REGION Network 9
   RUNG wire#powerrail
      { S7_Templates := "SrcType := Real" } LE_Contact(in1 := #"PID Output", in2 := #RangeY)
      Move(in := 0, out1 => #"Range2.Q")
   END_RUNG
   // the same network as SCL:
   IF #"PID Output" <= #RangeY THEN #"Range2.Q" := 0; END_IF;
END_REGION
END_FUNCTION_BLOCK

// folder: 1}Library/Timers

FUNCTION_BLOCK "TimerDisplay"   // FB2, LAD
{ S7_Optimized_Access := 'TRUE' }
VERSION : 0.1
   VAR_INPUT
      ET : DInt;
   END_VAR
   VAR_OUTPUT
      OUT : String;
   END_VAR
   VAR
      RealH : Real;
      RealM : Real;
      RealS : Real;
      RealMS : Real;
      StringH : String;
      StringM : String;
      StringS : String;
      StringMS : String;
      intH : Int;
      intM : Int;
      intS : Int;
      intMS : Int;
      String5 : String;
      String6 : String;
      String7 : String;
      String8 : String;
   END_VAR
   VAR_TEMP
      "dint-tempH" : DInt;
      "dint-tempM" : DInt;
      "dint-tempS" : DInt;
      "dint-tempMS" : DInt;
      "real-tempH" : Real;
      "real-tempM" : Real;
      "real-tempS" : Real;
      "real-tempMS" : Real;
   END_VAR
BEGIN

REGION Network 1: Reminder of H/M/S/MS
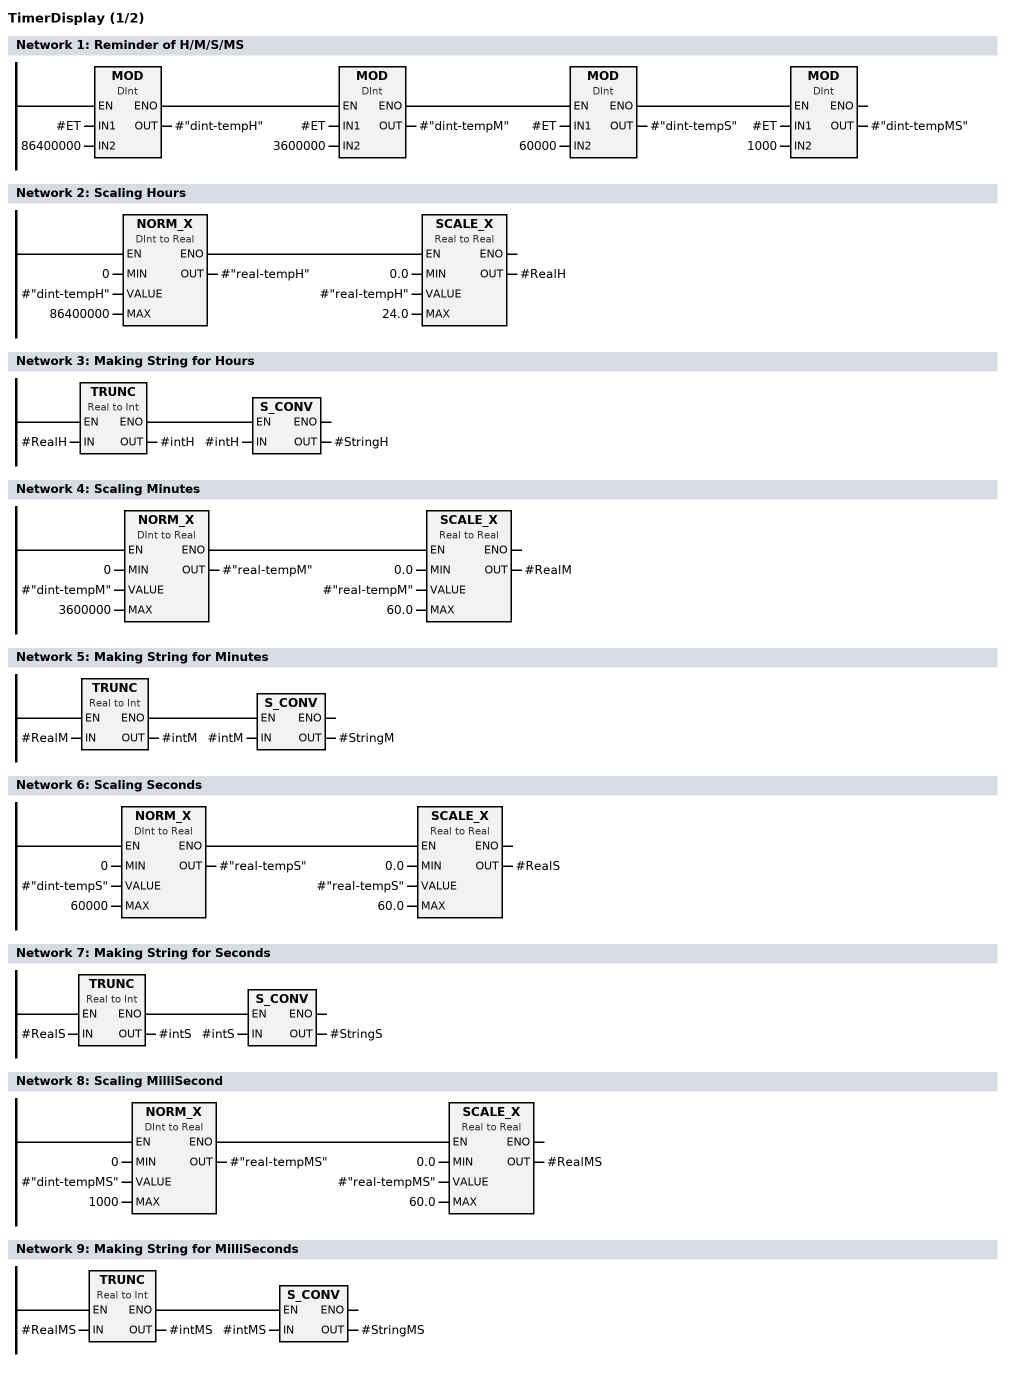
   RUNG wire#powerrail
      { S7_Templates := "SrcType := DInt" } Mod(in1 := #ET, in2 := 86400000, out => #"dint-tempH")
      { S7_Templates := "SrcType := DInt" } Mod(in1 := #ET, in2 := 3600000, out => #"dint-tempM")
      { S7_Templates := "SrcType := DInt" } Mod(in1 := #ET, in2 := 60000, out => #"dint-tempS")
      { S7_Templates := "SrcType := DInt" } Mod(in1 := #ET, in2 := 1000, out => #"dint-tempMS")
   END_RUNG
   // the same network as SCL:
   #"dint-tempH" := #ET MOD 86400000;
   #"dint-tempM" := #ET MOD 3600000;
   #"dint-tempS" := #ET MOD 60000;
   #"dint-tempMS" := #ET MOD 1000;
END_REGION

REGION Network 2: Scaling Hours
   RUNG wire#powerrail
      { S7_Templates := "[SrcType := DInt, DestType := Real]" } Normalize(min := 0, value := #"dint-tempH", max := 86400000, out => #"real-tempH")
      { S7_Templates := "[SrcType := Real, DestType := Real]" } Scale(min := 0.0, value := #"real-tempH", max := 24.0, out => #RealH)
   END_RUNG
   // the same network as SCL:
   #"real-tempH" := NORM_X(MIN := 0, VALUE := #"dint-tempH", MAX := 86400000);
   #RealH := SCALE_X(MIN := 0.0, VALUE := #"real-tempH", MAX := 24.0);
END_REGION

REGION Network 3: Making String for Hours
   #intH := TRUNC(#RealH);
   #StringH := S_CONV(IN := #intH);
END_REGION

REGION Network 4: Scaling Minutes
   RUNG wire#powerrail
      { S7_Templates := "[SrcType := DInt, DestType := Real]" } Normalize(min := 0, value := #"dint-tempM", max := 3600000, out => #"real-tempM")
      { S7_Templates := "[SrcType := Real, DestType := Real]" } Scale(min := 0.0, value := #"real-tempM", max := 60.0, out => #RealM)
   END_RUNG
   // the same network as SCL:
   #"real-tempM" := NORM_X(MIN := 0, VALUE := #"dint-tempM", MAX := 3600000);
   #RealM := SCALE_X(MIN := 0.0, VALUE := #"real-tempM", MAX := 60.0);
END_REGION

REGION Network 5: Making String for Minutes
   #intM := TRUNC(#RealM);
   #StringM := S_CONV(IN := #intM);
END_REGION

REGION Network 6: Scaling Seconds
   RUNG wire#powerrail
      { S7_Templates := "[SrcType := DInt, DestType := Real]" } Normalize(min := 0, value := #"dint-tempS", max := 60000, out => #"real-tempS")
      { S7_Templates := "[SrcType := Real, DestType := Real]" } Scale(min := 0.0, value := #"real-tempS", max := 60.0, out => #RealS)
   END_RUNG
   // the same network as SCL:
   #"real-tempS" := NORM_X(MIN := 0, VALUE := #"dint-tempS", MAX := 60000);
   #RealS := SCALE_X(MIN := 0.0, VALUE := #"real-tempS", MAX := 60.0);
END_REGION

REGION Network 7: Making String for Seconds
   #intS := TRUNC(#RealS);
   #StringS := S_CONV(IN := #intS);
END_REGION

REGION Network 8: Scaling MilliSecond
   RUNG wire#powerrail
      { S7_Templates := "[SrcType := DInt, DestType := Real]" } Normalize(min := 0, value := #"dint-tempMS", max := 1000, out => #"real-tempMS")
      { S7_Templates := "[SrcType := Real, DestType := Real]" } Scale(min := 0.0, value := #"real-tempMS", max := 60.0, out => #RealMS)
   END_RUNG
   // the same network as SCL:
   #"real-tempMS" := NORM_X(MIN := 0, VALUE := #"dint-tempMS", MAX := 1000);
   #RealMS := SCALE_X(MIN := 0.0, VALUE := #"real-tempMS", MAX := 60.0);
END_REGION

REGION Network 9: Making String for MilliSeconds
   #intMS := TRUNC(#RealMS);
   #StringMS := S_CONV(IN := #intMS);
END_REGION

REGION Network 10
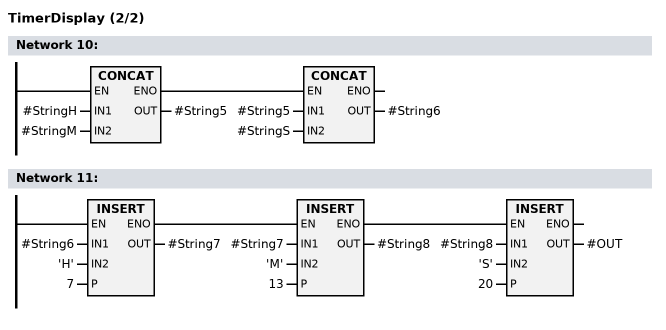
   #String5 := CONCAT(IN1 := #StringH, IN2 := #StringM);
   #String6 := CONCAT(IN1 := #String5, IN2 := #StringS);
END_REGION

REGION Network 11
   #String7 := INSERT(IN1 := #String6, IN2 := 'H', P := 7);
   #String8 := INSERT(IN1 := #String7, IN2 := 'M', P := 13);
   #OUT := INSERT(IN1 := #String8, IN2 := 'S', P := 20);
END_REGION
END_FUNCTION_BLOCK

// folder: 1}Library/Totalizer

FUNCTION_BLOCK "Totalizer_1"   // FB11, LAD
{ S7_Optimized_Access := 'TRUE' }
VERSION : 0.1
   VAR_INPUT
      value : Real;
      interval : Time;
      reset : Bool;
      cycle : Time;
   END_VAR
   VAR_OUTPUT
      Total : Real;
   END_VAR
   VAR
      accum1 : Real;
      accum2 : Real;
      "Timer" : IEC_TIMER;
   END_VAR
   VAR_TEMP
      tempInterval_Real : Real;
      tempInterval_Dint : DInt;
      tempCycle_Real : Real;
      tempCycle_Dint : Real;
      TempCalOne : Real;
      TempCalTwo : Real;
   END_VAR
BEGIN

REGION Network 1 (SCL): Reset Totalizer counts
   IF #reset THEN
       #accum1 := 0.0;
       #accum2 := 0.0;
       RESET_TIMER(#Timer);

   END_IF;
END_REGION

REGION Network 2 (SCL): Convert time into REAL
   #tempInterval_Real := TIME_TO_DINT (#interval);
   #tempCycle_Real := TIME_TO_DINT(#cycle);
END_REGION

REGION Network 3: Calculations for accum1
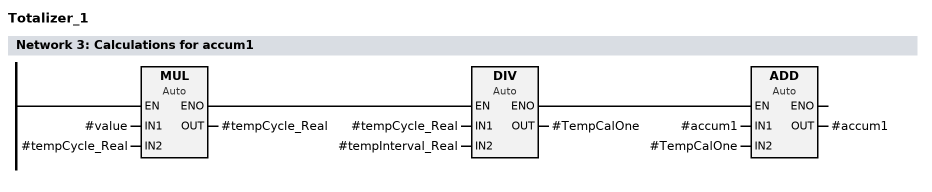
   RUNG wire#powerrail
      Mul(in1 := #value, in2 := #tempCycle_Real, out => #tempCycle_Real)
      Div(in1 := #tempCycle_Real, in2 := #tempInterval_Real, out => #TempCalOne)
      Add(in1 := #accum1, in2 := #TempCalOne, out => #accum1)
   END_RUNG
   // the same network as SCL:
   #tempCycle_Real := #value * #tempCycle_Real;
   #TempCalOne := #tempCycle_Real / #tempInterval_Real;
   #accum1 := #accum1 + #TempCalOne;
END_REGION

REGION Network 4 (SCL): Add the counters and reinitialize accum1
   IF #accum1 >= 1000.0 THEN
       #accum2 := 1000.0 + #accum2;
       #accum1 := 0.0;
   END_IF;

   #Total := #accum1 + #accum2;
END_REGION
END_FUNCTION_BLOCK

FUNCTION_BLOCK "Totalizer"   // FB17, LAD
{ S7_Optimized_Access := 'TRUE' }
VERSION : 0.1
   VAR_INPUT
      value : Real;
      interval : Time;
      reset : Bool;
      cycle : Time;
   END_VAR
   VAR_OUTPUT
      Total : Real;
   END_VAR
   VAR
      accum1 : Real;
      accum2 : Real;
      "Timer" : IEC_TIMER;
   END_VAR
   VAR_TEMP
      tempInterval_Real : Real;
      tempInterval_Dint : DInt;
      tempCycle_Real : Real;
      tempCycle_Dint : Real;
      TempCalOne : Real;
      TempCalTwo : Real;
   END_VAR
BEGIN

REGION Network 1 (SCL): Reset Totalizer counts
   IF #reset THEN
       #accum1 := 0.0;
       #accum2 := 0.0;
       #Total := 0.0;
       RESET_TIMER(#Timer);

   END_IF;
END_REGION

REGION Network 2 (SCL): Convert time into REAL
   #tempInterval_Real := TIME_TO_DINT (#interval);
   #tempCycle_Real := TIME_TO_DINT(#cycle);
END_REGION

REGION Network 3: Calculations for accum1
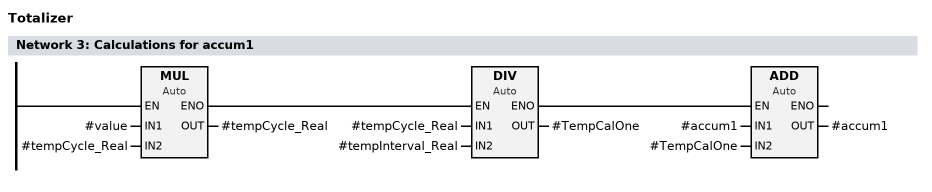
   RUNG wire#powerrail
      Mul(in1 := #value, in2 := #tempCycle_Real, out => #tempCycle_Real)
      Div(in1 := #tempCycle_Real, in2 := #tempInterval_Real, out => #TempCalOne)
      Add(in1 := #accum1, in2 := #TempCalOne, out => #accum1)
   END_RUNG
   // the same network as SCL:
   #tempCycle_Real := #value * #tempCycle_Real;
   #TempCalOne := #tempCycle_Real / #tempInterval_Real;
   #accum1 := #accum1 + #TempCalOne;
END_REGION

REGION Network 4 (SCL): Add the counters and reinitialize accum1
   IF #accum1 >= 1000.0 THEN
       #accum2 := 1000.0 + #accum2;
       #accum1 := 0.0;
   END_IF;

   #Total := #accum1 + #accum2;
END_REGION
END_FUNCTION_BLOCK

// folder: 1}Library/VFD

FUNCTION_BLOCK "VFD_PNCtrl"   // FB9, SCL
TITLE = VFD Controlled by Profinet
{ S7_Optimized_Access := 'TRUE' }
VERSION : 0.1
   VAR_INPUT
      EnableBlock : Bool;
      EnableAxis : Bool;
      AckError : Bool;
      SpeedSP_Perc : Real;   // Speed SP in Percentage 0-100%
      RefSpeed : Real;   // Reference Speed in RPM (parameter p2000)
      ConfigAxis : Word := 16#003F;
      HWIDSTW : Hw_Io;
      HWIDZSW : Hw_Io;
   END_VAR
   VAR_OUTPUT
      AxisEnabled : Bool;
      Lockout : Bool;
      ActVelocity_Perc : Real;
      ActVelocity_RPM : Real;
      Error : Bool;
      Status : Word;
      DiagId : Word;
   END_VAR
   VAR
      SP_Rpm : Real;   // Speed SP in RPM
      SinaSpeed_Instance : SinaSpeed;
   END_VAR
BEGIN
   //******************************************************************************
   //Convert Speed SP from Percentage to RPM

   #SP_Rpm := (#SpeedSP_Perc * #RefSpeed) / 100;

   IF #EnableBlock THEN


       #SinaSpeed_Instance(EnableAxis := #EnableAxis,
                           AckError := #AckError,
                           SpeedSp := #SP_Rpm,
                           RefSpeed := #RefSpeed,
                           ConfigAxis := #ConfigAxis,
                           HWIDSTW := #HWIDSTW,
                           HWIDZSW := #HWIDZSW,
                           AxisEnabled => #AxisEnabled,
                           Lockout => #Lockout,
                           ActVelocity => #ActVelocity_Perc,
                           Error => #Error,
                           Status => #Status,
                           DiagId => #DiagId);

   ELSE

       #SinaSpeed_Instance(EnableAxis := FALSE,
                           AckError :=FALSE,
                           SpeedSp := 0.0,
                           RefSpeed := #RefSpeed,
                           ConfigAxis := #ConfigAxis,
                           HWIDSTW := #HWIDSTW,
                           HWIDZSW := #HWIDZSW,
                           AxisEnabled => #AxisEnabled,
                           Lockout => #Lockout,
                           ActVelocity => #ActVelocity_Perc,
                           Error => #Error,
                           Status => #Status,
                           DiagId => #DiagId);


       #Error := FALSE;

   END_IF;

   #ActVelocity_Perc := (#SinaSpeed_Instance.ActVelocity * 100) / #RefSpeed;
   #ActVelocity_RPM := #SinaSpeed_Instance.ActVelocity;
END_FUNCTION_BLOCK

FUNCTION_BLOCK "VFD_Dumbdown"   // FB812, LAD
{ S7_Optimized_Access := 'TRUE' }
VERSION : 0.7
   VAR_INPUT
      IL : Bool := TRUE;   // Interlock
      PLCCommand : Bool;   // Auto Command to Run (logic from PLC to command motor to run)
      RUN_FEEDBACK : Bool;   // Feedback from the drive indicating that it is running
      VFD_FAULT : Bool;   // Feedback from the drive that it is in Fault
      AUTO_SPEED_P : Word;   // Auto Speed Setpoint Command (logic from PLC to command motor speed) Raw 0-27648
      AUTO_SPEED_R : Real;   // Auto Speed Setpoint Command (logic from PLC to command motor speed) Scale 0-100
      SPEED_FEEDBACK : Int;   // Speed Feedback raw Siganl from the drive
   END_VAR
   VAR_OUTPUT
      RUN_CMD : Bool;
      Stop_CMD : Bool;   // Stop Command
      Start_CMD : Bool;   // Start Command
      RST_CMD : Bool;   // VFD Reset
      VFD_SPEED : Int;   // Command Speed Setpoint to VFD
      VFD_TORQUE : Int;   // Command Torque Setpoint to VFD
   END_VAR
   VAR
      HMI : Struct   // Struct for HMI
         Controls : Struct
            Mode : Int;   // HOA = Auto, 0 = Off, 1 = Manual (HMI Control), 2 = Auto (PLC Control)
            Start : Bool;   // Mode = 1, Start VFD Command
            Stop : Bool;   // Mode = 1, Stop VFD Command
            Reset : Bool;   // VFD Reset Command
            PLCMOHR : Bool;   // PLC Motor Operating Hours Reset
            Speed_Setpoint : Real;   // Speed Setpoint to Drive Real 0-100.0
         END_STRUCT;
         Status : Struct
            HOAStatus : Int;   // HOA Status
            PLC_MOH : Real;
            LMOH : Real;   // Last Motor Operating Hours
            VFDON : Bool;   // VFD On
            VFD_FAULT : Bool;   // VFD is Faulted
            CMD : Bool;   // Commanding VFD to Run
            IL : Bool;   // Interlock Active
            VFD_SPEED : Real;   // VFD Speed Feedback from the drive
            VFD_TORQUE : Real;
         END_STRUCT;
         Config : Struct
            RCPD_SP : Int := 300;
            Start_PT : Time := T#500MS;
            Stop_PT : Time := T#500MS;
         END_STRUCT;
      END_STRUCT;
      Math : Struct
         MOH1 : DInt;
         MOH2 : Real;
         PLCMOH : Real;   // PLC Motor Operating Hours
         LMOH : Real;
      END_STRUCT;
      OS : Struct
         RON : Bool;   // Remote / HMI On
         ROFF : Bool;   // Remote / HMI Off
         HON : Bool;   // Hand/Local On
         Auto : Bool;   // Auto
         PLCMOHR : Bool;
         LMOH1 : Bool;
         LMOH2 : Bool;
         RST : Bool;   // Reset VFD
         Bipolar : Bool;
         MinuteTime : Bool;
         HoursTime : Real;
         Raw_Auto_Speed_Set : Int;
         Unscale_Return : Word;
      END_STRUCT;
      Motor_max_RPM : Real := 100.0;
      START_CMD_TOF : IEC_TIMER;   // Start Semicode
      STOP_CMD_TOF : IEC_TIMER;
      Reset_Hold_Time : IEC_TIMER;
      Motor_Minute_Counter : IEC_TIMER;
      TIMEOUT : IEC_TIMER;
   END_VAR
   VAR_TEMP   // added for the SCL form of the ladder/FBD networks
      _w1 : Bool;
      _w2 : Bool;
   END_VAR
BEGIN

REGION Network 1: Start VFD
   // Main Logic of the FB
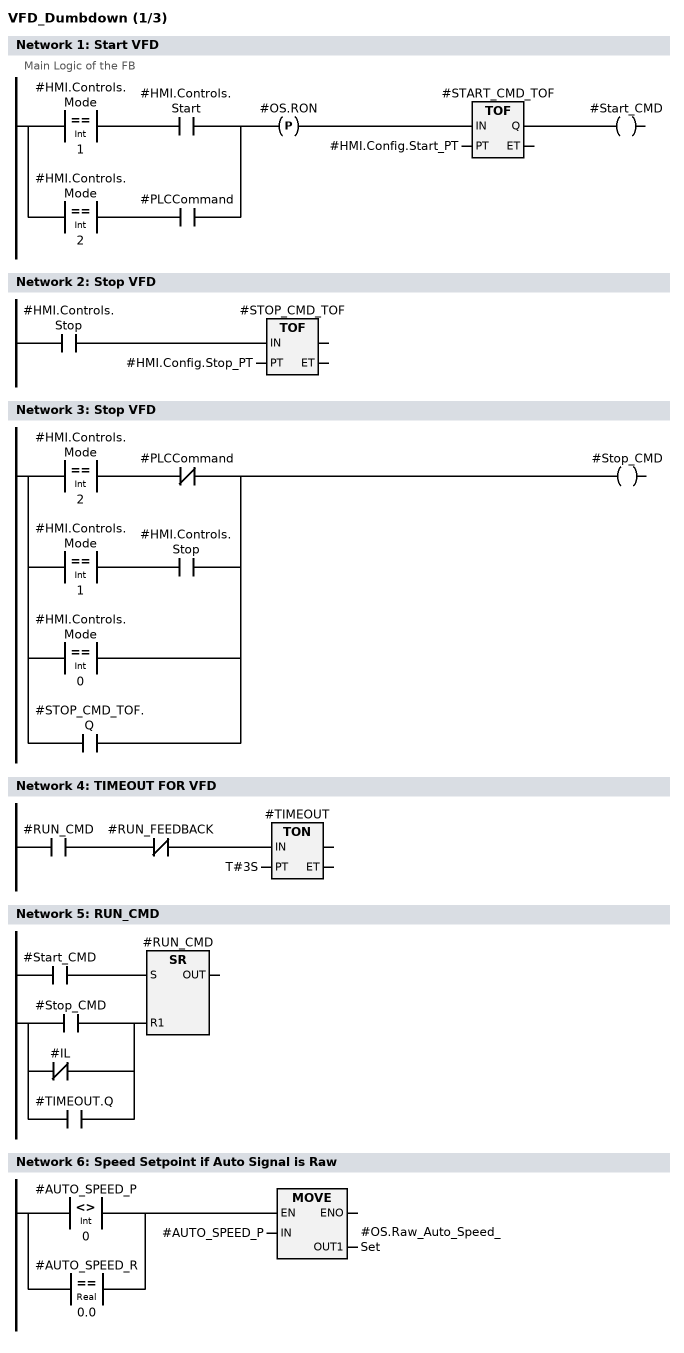
   #_w1 := ((#HMI.Controls.Mode = 1) AND #HMI.Controls.Start) OR ((#HMI.Controls.Mode = 2) AND #PLCCommand);
   #_w2 := #_w1 AND NOT #OS.RON;   // rising edge
   #OS.RON := #_w1;
   #START_CMD_TOF.TOF(IN := #_w2, PT := #HMI.Config.Start_PT);
   #Start_CMD := #START_CMD_TOF.Q;
END_REGION

REGION Network 2: Stop VFD
   #STOP_CMD_TOF.TOF(IN := #HMI.Controls.Stop, PT := #HMI.Config.Stop_PT);
END_REGION

REGION Network 3: Stop VFD
   RUNG wire#powerrail
      { S7_Templates := "SrcType := Int" } EQ_Contact(in1 := #HMI.Controls.Mode, in2 := 2)
      I_Contact( #PLCCommand )
      wire#w1
      Coil( #Stop_CMD )
   END_RUNG
   RUNG wire#powerrail
      { S7_Templates := "SrcType := Int" } EQ_Contact(in1 := #HMI.Controls.Mode, in2 := 1)
      Contact( #HMI.Controls.Stop )
   END_RUNG wire#w1
   RUNG wire#powerrail
      { S7_Templates := "SrcType := Int" } EQ_Contact(in1 := #HMI.Controls.Mode, in2 := 0)
   END_RUNG wire#w1
   RUNG wire#powerrail
      Contact( #STOP_CMD_TOF.Q )
   END_RUNG wire#w1
   // the same network as SCL:
   #Stop_CMD := ((#HMI.Controls.Mode = 2) AND NOT #PLCCommand) OR ((#HMI.Controls.Mode = 1) AND #HMI.Controls.Stop) OR (#HMI.Controls.Mode = 0) OR #STOP_CMD_TOF.Q;
END_REGION

REGION Network 4: TIMEOUT FOR VFD
   #TIMEOUT.TON(IN := #RUN_CMD AND NOT #RUN_FEEDBACK, PT := T#3S);
END_REGION

REGION Network 5: RUN_CMD
   RUNG wire#powerrail
      Contact( #Start_CMD )
      S_SR(operand := #RUN_CMD, r1 := wire#w1)
   END_RUNG
   RUNG wire#powerrail
      Contact( #Stop_CMD )
   END_RUNG wire#w1
   RUNG wire#powerrail
      I_Contact( #IL )
   END_RUNG wire#w1
   RUNG wire#powerrail
      Contact( #TIMEOUT.Q )
   END_RUNG wire#w1
   // the same network as SCL:
   IF #Start_CMD THEN
       #RUN_CMD := TRUE;   // SR flip-flop
   END_IF;
   IF #Stop_CMD OR NOT #IL OR #TIMEOUT.Q THEN #RUN_CMD := FALSE; END_IF;
END_REGION

REGION Network 6: Speed Setpoint if Auto Signal is Raw
   RUNG wire#powerrail
      { S7_Templates := "SrcType := Int" } NE_Contact(in1 := #AUTO_SPEED_P, in2 := 0)
      wire#w1
      { S7_GenerateENO := "TRUE" } Move(in := #AUTO_SPEED_P, out1 => #OS.Raw_Auto_Speed_Set)
   END_RUNG
   RUNG wire#powerrail
      { S7_Templates := "SrcType := Real" } EQ_Contact(in1 := #AUTO_SPEED_R, in2 := 0.0)
   END_RUNG wire#w1
   // the same network as SCL:
   IF (#AUTO_SPEED_P <> 0) OR (#AUTO_SPEED_R = 0.0) THEN #OS.Raw_Auto_Speed_Set := #AUTO_SPEED_P; END_IF;
END_REGION

REGION Network 7: Speed Setpoint if Auto Signal is Real
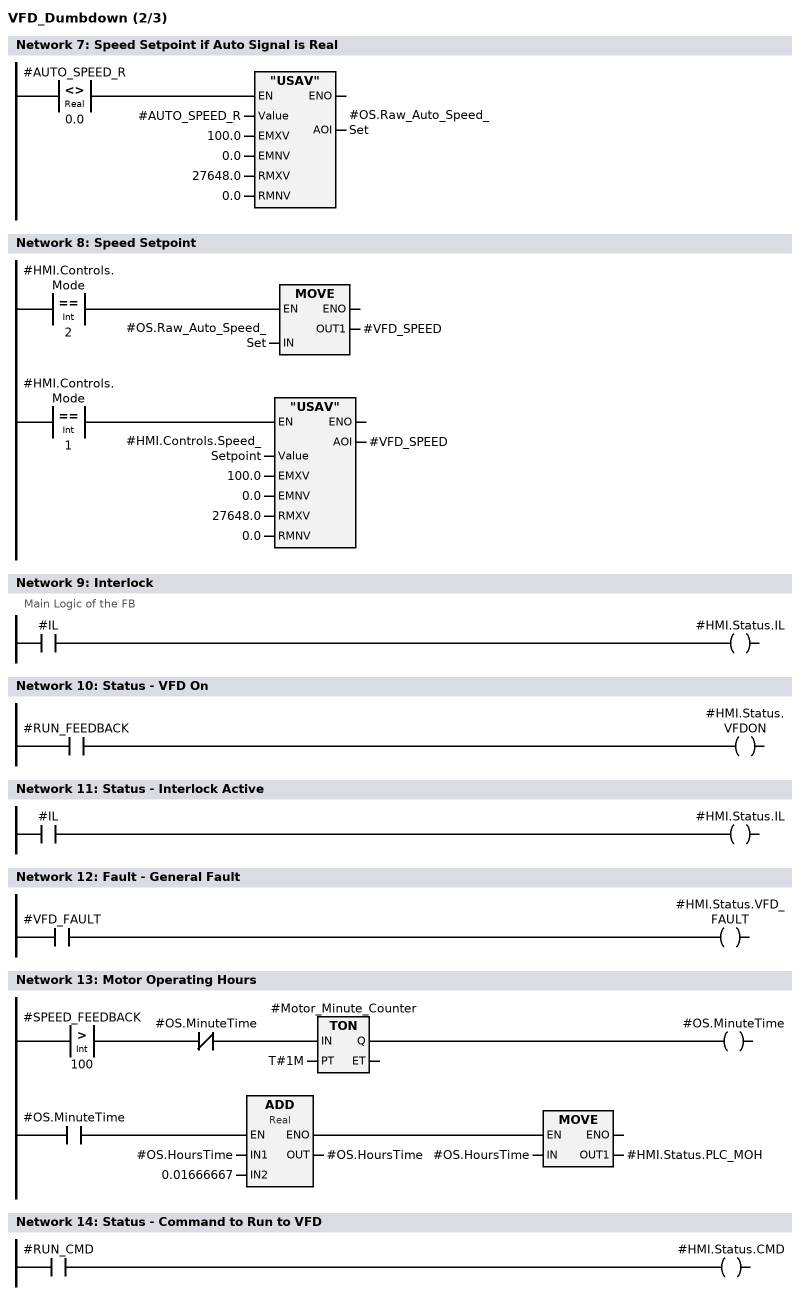
   RUNG wire#powerrail
      { S7_Templates := "SrcType := Real" } NE_Contact(in1 := #AUTO_SPEED_R, in2 := 0.0)
      "USAV"(Value := #AUTO_SPEED_R, EMXV := 100.0, EMNV := 0.0, RMXV := 27648.0, RMNV := 0.0, AOI => #OS.Raw_Auto_Speed_Set)
   END_RUNG
   // the same network as SCL:
   IF #AUTO_SPEED_R <> 0.0 THEN
       "USAV"(Value := #AUTO_SPEED_R,
              EMXV := 100.0,
              EMNV := 0.0,
              RMXV := 27648.0,
              RMNV := 0.0,
              AOI => #OS.Raw_Auto_Speed_Set);
   END_IF;
END_REGION

REGION Network 8: Speed Setpoint
   RUNG wire#powerrail
      { S7_Templates := "SrcType := Int" } EQ_Contact(in1 := #HMI.Controls.Mode, in2 := 2)
      { S7_GenerateENO := "TRUE" } Move(in := #OS.Raw_Auto_Speed_Set, out1 => #VFD_SPEED)
   END_RUNG
   RUNG wire#powerrail
      { S7_Templates := "SrcType := Int" } EQ_Contact(in1 := #HMI.Controls.Mode, in2 := 1)
      "USAV"(Value := #HMI.Controls.Speed_Setpoint, EMXV := 100.0, EMNV := 0.0, RMXV := 27648.0, RMNV := 0.0, AOI => #VFD_SPEED)
   END_RUNG
   // the same network as SCL:
   IF #HMI.Controls.Mode = 2 THEN #VFD_SPEED := #OS.Raw_Auto_Speed_Set; END_IF;
   IF #HMI.Controls.Mode = 1 THEN
       "USAV"(Value := #HMI.Controls.Speed_Setpoint,
              EMXV := 100.0,
              EMNV := 0.0,
              RMXV := 27648.0,
              RMNV := 0.0,
              AOI => #VFD_SPEED);
   END_IF;
END_REGION

REGION Network 9: Interlock
   // Main Logic of the FB
   RUNG wire#powerrail
      Contact( #IL )
      Coil( #HMI.Status.IL )
   END_RUNG
   // the same network as SCL:
   #HMI.Status.IL := #IL;
END_REGION

REGION Network 10: Status - VFD On
   RUNG wire#powerrail
      Contact( #RUN_FEEDBACK )
      Coil( #HMI.Status.VFDON )
   END_RUNG
   // the same network as SCL:
   #HMI.Status.VFDON := #RUN_FEEDBACK;
END_REGION

REGION Network 11: Status - Interlock Active
   RUNG wire#powerrail
      Contact( #IL )
      Coil( #HMI.Status.IL )
   END_RUNG
   // the same network as SCL:
   #HMI.Status.IL := #IL;
END_REGION

REGION Network 12: Fault - General Fault
   RUNG wire#powerrail
      Contact( #VFD_FAULT )
      Coil( #HMI.Status.VFD_FAULT )
   END_RUNG
   // the same network as SCL:
   #HMI.Status.VFD_FAULT := #VFD_FAULT;
END_REGION

REGION Network 13: Motor Operating Hours
   #Motor_Minute_Counter.TON(IN := (#SPEED_FEEDBACK > 100) AND NOT #OS.MinuteTime, PT := T#1M);
   #OS.MinuteTime := #Motor_Minute_Counter.Q;
   IF #OS.MinuteTime THEN
       #OS.HoursTime := #OS.HoursTime + 0.01666667;
       #HMI.Status.PLC_MOH := #OS.HoursTime;
   END_IF;
END_REGION

REGION Network 14: Status - Command to Run to VFD
   RUNG wire#powerrail
      Contact( #RUN_CMD )
      Coil( #HMI.Status.CMD )
   END_RUNG
   // the same network as SCL:
   #HMI.Status.CMD := #RUN_CMD;
END_REGION

REGION Network 15: VFD Speed Feedback
   // VFD Speed Feedback
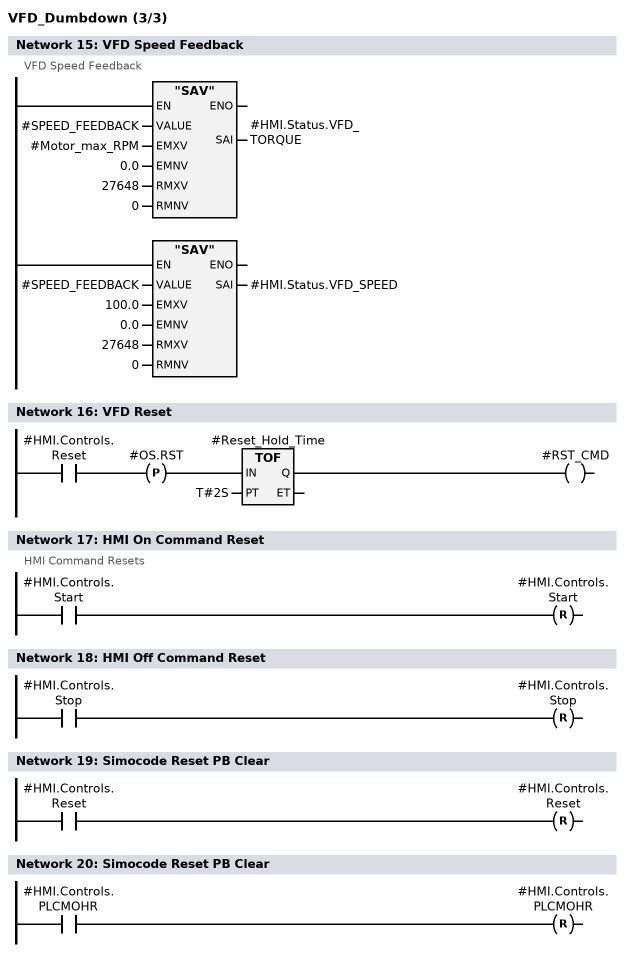
   RUNG wire#powerrail
      "SAV"(VALUE := #SPEED_FEEDBACK, EMXV := #Motor_max_RPM, EMNV := 0.0, RMXV := 27648, RMNV := 0, SAI => #HMI.Status.VFD_TORQUE)
   END_RUNG
   RUNG wire#powerrail
      "SAV"(VALUE := #SPEED_FEEDBACK, EMXV := 100.0, EMNV := 0.0, RMXV := 27648, RMNV := 0, SAI => #HMI.Status.VFD_SPEED)
   END_RUNG
   // the same network as SCL:
   "SAV"(VALUE := #SPEED_FEEDBACK,
         EMXV := #Motor_max_RPM,
         EMNV := 0.0,
         RMXV := 27648,
         RMNV := 0,
         SAI => #HMI.Status.VFD_TORQUE);
   "SAV"(VALUE := #SPEED_FEEDBACK,
         EMXV := 100.0,
         EMNV := 0.0,
         RMXV := 27648,
         RMNV := 0,
         SAI => #HMI.Status.VFD_SPEED);
END_REGION

REGION Network 16: VFD Reset
   #_w1 := #HMI.Controls.Reset AND NOT #OS.RST;   // rising edge
   #OS.RST := #HMI.Controls.Reset;
   #Reset_Hold_Time.TOF(IN := #_w1, PT := T#2S);
   #RST_CMD := #Reset_Hold_Time.Q;
END_REGION

REGION Network 17: HMI On Command Reset
   // HMI Command Resets
   RUNG wire#powerrail
      Contact( #HMI.Controls.Start )
      R_Coil( #HMI.Controls.Start )
   END_RUNG
   // the same network as SCL:
   IF #HMI.Controls.Start THEN #HMI.Controls.Start := FALSE; END_IF;
END_REGION

REGION Network 18: HMI Off Command Reset
   RUNG wire#powerrail
      Contact( #HMI.Controls.Stop )
      R_Coil( #HMI.Controls.Stop )
   END_RUNG
   // the same network as SCL:
   IF #HMI.Controls.Stop THEN #HMI.Controls.Stop := FALSE; END_IF;
END_REGION

REGION Network 19: Simocode Reset PB Clear
   RUNG wire#powerrail
      Contact( #HMI.Controls.Reset )
      R_Coil( #HMI.Controls.Reset )
   END_RUNG
   // the same network as SCL:
   IF #HMI.Controls.Reset THEN #HMI.Controls.Reset := FALSE; END_IF;
END_REGION

REGION Network 20: Simocode Reset PB Clear
   RUNG wire#powerrail
      Contact( #HMI.Controls.PLCMOHR )
      R_Coil( #HMI.Controls.PLCMOHR )
   END_RUNG
   // the same network as SCL:
   IF #HMI.Controls.PLCMOHR THEN #HMI.Controls.PLCMOHR := FALSE; END_IF;
END_REGION
END_FUNCTION_BLOCK

// folder: 1}Library/Valve

FUNCTION_BLOCK "Valve-SV"   // FB800, LAD
{ S7_Optimized_Access := 'FALSE' }
VERSION : 1.0
   VAR_INPUT
      OS : Bool;   // Open Signal
      CS : Bool;   // Close Signal
      VML : Bool;   // Valve Mode set to Local
      VMR : Bool := TRUE;   // Valve Mode set to Remote
      EI : Bool := TRUE;   // Indication - ESD
      EM : Int := 0;   // Mode - 0=FC / 1=FO / 2=FL
      CP : Bool := TRUE;   // Control - Permissive
      LOR : Bool;   // Local/Off/Remote indications are N/A
      MC : Bool := TRUE;   // Maintained Command
      VT : Int := 3;   // 0 = 2 In 2 Out // 1 = 1 In 2 Outs // 2 = 2 In 1 Out // 3 = 1 In 1 Out
   END_VAR
   VAR_OUTPUT
      AVL : Bool;   // Valve available to be remotely controlled
      CO : Bool;   // Command Open
      CC : Bool;   // Command Close
   END_VAR
   VAR
      CMD : Int;   // 0=Stop / 1=Close / 2=Open
      Lockout : Bool;
      Status : Struct
         CP : Int;   // Current Position = (0=Open) (1=In Transition) (2=Close) (3=No Position)
      END_STRUCT;
      Alarms : Struct
         "TO" : Bool;   // Alarm - Open Timeout
         TC : Bool;   // Alarm - Close Timeout
         TNOCR : Bool;   // Alarm - Total Number of Open Commands Reached
         TNCCR : Bool;   // Alarm - Total Number of Close Commands Reached
      END_STRUCT;
      Timeouts : Struct
         OTS : Time := t#30s;   // Open Timeout Setpoint
         CTS : Time := t#30s;   // Close Timeout Setpoint
      END_STRUCT;
      Pulse : Struct
         TOP : Bool;   // Timeout - Open pulse
         TCP : Bool;   // Timeout - Close pulse
         TOR : Bool;   // Timeout - Open Reset
         TCR : Bool;   // Timeout - Open Reset
         VOP : Bool;   // Verified Open Pulse
         VCP : Bool;   // Verified Close Pulse
         LCO : Bool;   // Last Command Open
         LCC : Bool;   // Last Command Close
         OSP : Bool;   // Open Status Pulse
         CSP : Bool;   // Close Status Pulse
         TSP : Bool;   // Transition Status Pulse
         NSP : Bool;   // No Status Position
      END_STRUCT;
      Save : Struct
         LC : Int;   // Last Command from Operator
         STOC : Int;   // Service Total Open Commands
         STCC : Int;   // Service Total Close Commands
         PS : Bool;   // Permissive Save
      END_STRUCT;
      Diags : Struct
         STOCS : Int := 9999;   // Service Total Open Commands Setpoint
         STCCS : Int := 9999;   // Service Total Close Commands Setpoint
      END_STRUCT;
      AVL_DBNC : TON_TIME;   // Valve Availability Debounce
      TO_O : TON_TIME;   // Timeout - Open
      TO_C : TON_TIME;   // Timeout - Close
      VRFD_O : TON_TIME;   // Verified - Successful open
      VRFD_C : TON_TIME;   // Verified - Successful close
      TSOC : CTU_INT;   // Total Service Open Commands
      TSCC : CTU_INT;   // Total Service Close Commands
      AVL_HLD_TOF : TOF_TIME;   // Valve Availability Hold
      Mode : Int := 1;   // Mode Man=1, Aut=0
   END_VAR
   VAR_TEMP
      VA : Bool;   // Valve Available
      TCO : Bool;   // Temp Command Open
      TCC : Bool;   // Temp Command Close
      TAVL : Bool;   // Temp Available
   END_VAR
   VAR_TEMP   // added for the SCL form of the ladder/FBD networks
      _w1 : Bool;
      _w2 : Bool;
      _w3 : Bool;
      _w4 : Bool;
   END_VAR
BEGIN

REGION Network 1: Function Block Mode = 0
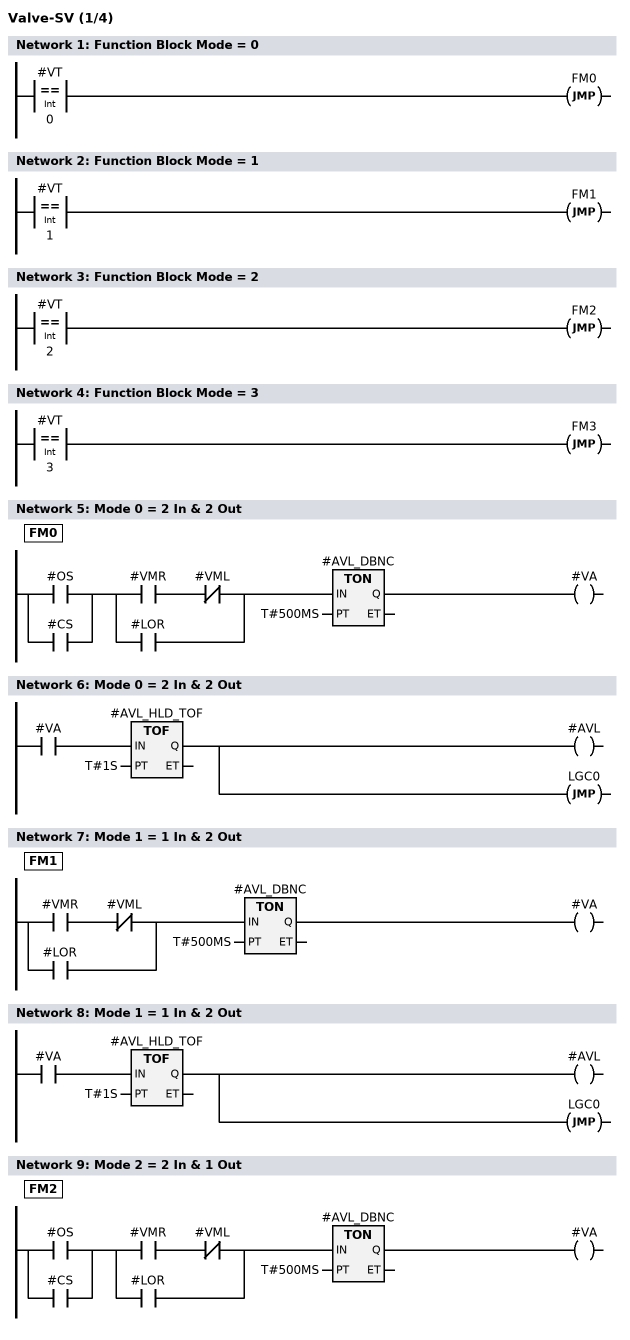
   RUNG wire#powerrail
      { S7_Templates := "SrcType := Int" } EQ_Contact(in1 := #VT, in2 := 0)
      JumpCoil( FM0 )
   END_RUNG
   // the same network as SCL:
   IF #VT = 0 THEN GOTO FM0; END_IF;
END_REGION

REGION Network 2: Function Block Mode = 1
   RUNG wire#powerrail
      { S7_Templates := "SrcType := Int" } EQ_Contact(in1 := #VT, in2 := 1)
      JumpCoil( FM1 )
   END_RUNG
   // the same network as SCL:
   IF #VT = 1 THEN GOTO FM1; END_IF;
END_REGION

REGION Network 3: Function Block Mode = 2
   RUNG wire#powerrail
      { S7_Templates := "SrcType := Int" } EQ_Contact(in1 := #VT, in2 := 2)
      JumpCoil( FM2 )
   END_RUNG
   // the same network as SCL:
   IF #VT = 2 THEN GOTO FM2; END_IF;
END_REGION

REGION Network 4: Function Block Mode = 3
   RUNG wire#powerrail
      { S7_Templates := "SrcType := Int" } EQ_Contact(in1 := #VT, in2 := 3)
      JumpCoil( FM3 )
   END_RUNG
   // the same network as SCL:
   IF #VT = 3 THEN GOTO FM3; END_IF;
END_REGION

REGION Network 5: Mode 0 = 2 In & 2 Out
   FM0:
   #AVL_DBNC(IN := (#OS OR #CS) AND ((#VMR AND NOT #VML) OR #LOR), PT := T#500MS);   // TON
   #VA := #AVL_DBNC.Q;
END_REGION

REGION Network 6: Mode 0 = 2 In & 2 Out
   #AVL_HLD_TOF(IN := #VA, PT := T#1S);   // TOF
   #AVL := #AVL_HLD_TOF.Q;
   IF #AVL_HLD_TOF.Q THEN GOTO LGC0; END_IF;
END_REGION

REGION Network 7: Mode 1 = 1 In & 2 Out
   FM1:
   #AVL_DBNC(IN := (#VMR AND NOT #VML) OR #LOR, PT := T#500MS);   // TON
   #VA := #AVL_DBNC.Q;
END_REGION

REGION Network 8: Mode 1 = 1 In & 2 Out
   #AVL_HLD_TOF(IN := #VA, PT := T#1S);   // TOF
   #AVL := #AVL_HLD_TOF.Q;
   IF #AVL_HLD_TOF.Q THEN GOTO LGC0; END_IF;
END_REGION

REGION Network 9: Mode 2 = 2 In & 1 Out
   FM2:
   #AVL_DBNC(IN := (#OS OR #CS) AND ((#VMR AND NOT #VML) OR #LOR), PT := T#500MS);   // TON
   #VA := #AVL_DBNC.Q;
END_REGION

REGION Network 10: Mode 2 = 2 In & 1 Out
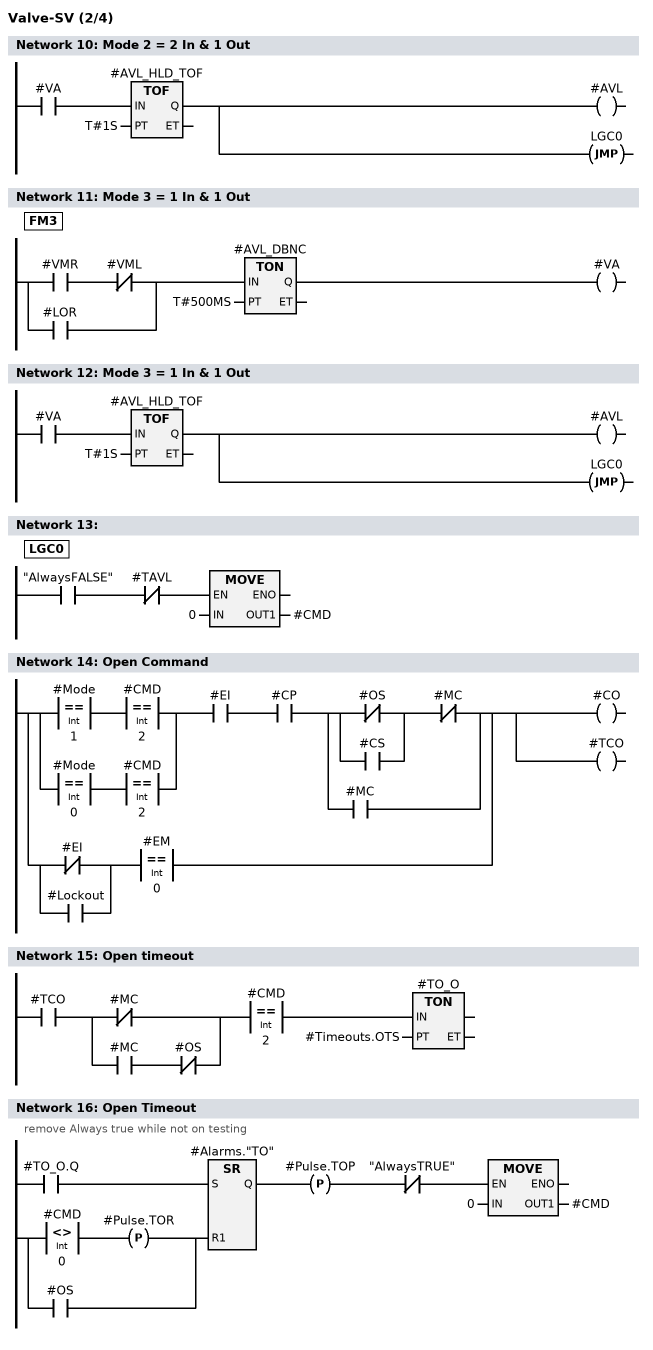
   #AVL_HLD_TOF(IN := #VA, PT := T#1S);   // TOF
   #AVL := #AVL_HLD_TOF.Q;
   IF #AVL_HLD_TOF.Q THEN GOTO LGC0; END_IF;
END_REGION

REGION Network 11: Mode 3 = 1 In & 1 Out
   FM3:
   #AVL_DBNC(IN := (#VMR AND NOT #VML) OR #LOR, PT := T#500MS);   // TON
   #VA := #AVL_DBNC.Q;
END_REGION

REGION Network 12: Mode 3 = 1 In & 1 Out
   #AVL_HLD_TOF(IN := #VA, PT := T#1S);   // TOF
   #AVL := #AVL_HLD_TOF.Q;
   IF #AVL_HLD_TOF.Q THEN GOTO LGC0; END_IF;
END_REGION

REGION Network 13
   Label( LGC0 )
   RUNG wire#powerrail
      Contact( "AlwaysFALSE" )
      I_Contact( #TAVL )
      { S7_GenerateENO := "TRUE" } Move(in := 0, out1 => #CMD)
   END_RUNG
   // the same network as SCL:
   LGC0:
   IF "AlwaysFALSE" AND NOT #TAVL THEN #CMD := 0; END_IF;
END_REGION

REGION Network 14: Open Command
   RUNG wire#powerrail
      { S7_Templates := "SrcType := Int" } EQ_Contact(in1 := #Mode, in2 := 1)
      { S7_Templates := "SrcType := Int" } EQ_Contact(in1 := #CMD, in2 := 2)
      wire#w1
      Contact( #EI )
      Contact( #CP )
      wire#w2
      I_Contact( #OS )
      wire#w3
      I_Contact( #MC )
      wire#w4
      Coil( #CO )
   END_RUNG
   RUNG wire#powerrail
      { S7_Templates := "SrcType := Int" } EQ_Contact(in1 := #Mode, in2 := 0)
      { S7_Templates := "SrcType := Int" } EQ_Contact(in1 := #CMD, in2 := 2)
   END_RUNG wire#w1
   RUNG wire#w2
      Contact( #CS )
   END_RUNG wire#w3
   RUNG wire#w2
      Contact( #MC )
   END_RUNG wire#w4
   RUNG wire#powerrail
      I_Contact( #EI )
      wire#w5
      { S7_Templates := "SrcType := Int" } EQ_Contact(in1 := #EM, in2 := 0)
   END_RUNG wire#w4
   RUNG wire#powerrail
      Contact( #Lockout )
   END_RUNG wire#w5
   RUNG wire#w4
      Coil( #TCO )
   END_RUNG
   // the same network as SCL:
   #CO := ((((#Mode = 1) AND (#CMD = 2)) OR ((#Mode = 0) AND (#CMD = 2))) AND #EI AND #CP AND (((NOT #OS OR #CS) AND NOT #MC) OR #MC)) OR ((NOT #EI OR #Lockout) AND (#EM = 0));
   #TCO := #CO;
END_REGION

REGION Network 15: Open timeout
   #TO_O(IN := #TCO AND (NOT #MC OR (#MC AND NOT #OS)) AND (#CMD = 2), PT := #Timeouts.OTS);   // TON
END_REGION

REGION Network 16: Open Timeout
   // remove Always true while not on testing
   RUNG wire#powerrail
      Contact( #TO_O.Q )
      S_SR(operand := #Alarms."TO", r1 := wire#w1)
      P_Trig( #Pulse.TOP )
      I_Contact( "AlwaysTRUE" )
      { S7_GenerateENO := "TRUE" } Move(in := 0, out1 => #CMD)
   END_RUNG
   RUNG wire#powerrail
      { S7_Templates := "SrcType := Int" } NE_Contact(in1 := #CMD, in2 := 0)
      P_Trig( #Pulse.TOR )
   END_RUNG wire#w1
   RUNG wire#powerrail
      Contact( #OS )
   END_RUNG wire#w1
   // the same network as SCL:
   #_w1 := #CMD <> 0;
   #_w2 := #_w1 AND NOT #Pulse.TOR;   // rising edge
   #Pulse.TOR := #_w1;
   IF #TO_O.Q THEN
       #Alarms."TO" := TRUE;   // SR flip-flop
   END_IF;
   IF #_w2 OR #OS THEN #Alarms."TO" := FALSE; END_IF;
   #_w3 := #Alarms."TO" AND NOT #Pulse.TOP;   // rising edge
   #Pulse.TOP := #Alarms."TO";
   IF #_w3 AND NOT "AlwaysTRUE" THEN #CMD := 0; END_IF;
END_REGION

